VERSION : 0.1
   VAR_INPUT
      codeLib : "From Excel: Data";
   END_VAR
   VAR_IN_OUT
      savedWipStns : "Recipe: HMI Stations Saved Wips";
   END_VAR
   VAR_TEMP
      pStn : Int;
      pDestStn : Int;
      pWip : Int;
   END_VAR
BEGIN
   REGION "HMI STATIONS"
       FOR #pStn := 0 TO UDINT_TO_INT("Length"(#codeLib.hmiStns) - 1) DO
           #pDestStn := #codeLib.hmiStns[#pStn].pStn;
           IF #pDestStn = -1 THEN
               EXIT;
           END_IF;
           FOR #pWip := 0 TO "wipCount" DO
               #savedWipStns.stn[#pStn].wip[#pWip].pnCode :=
                   #codeLib.hmiStns[#pStn].wip[#pWip].pnCode;
           END_FOR;
       END_FOR;
   END_REGION
END_FUNCTION

FUNCTION "From Excel: PN Code to HMI Stations" : Void   // FC62, SCL
{ S7_Optimized_Access := 'TRUE' }
VERSION : 0.1
   VAR_INPUT
      xlCodeLib : "From Excel: Data";
   END_VAR
   VAR_IN_OUT
      stns : "Station: All Stations";
   END_VAR
   VAR_TEMP
      pSrc : Int;
      pDest : Int;
   END_VAR
BEGIN
   REGION "HMI STATIONS"
       FOR #pSrc := 0 TO UDINT_TO_INT("Length"(#xlCodeLib.hmiStns) - 1) DO
           #pDest := #xlCodeLib.hmiStns[#pSrc].pStn;
           IF #pDest = -1 THEN
               EXIT;
           END_IF;
           #stns.stn[#pDest].wipCmpts.pnCode := #xlCodeLib.hmiStns[#pSrc].wip[0].pnCode;
       END_FOR;
   END_REGION
END_FUNCTION

FUNCTION "From Excel: Wip Code to HMI Station Saved WIps" : Void   // FC63, SCL
{ S7_Optimized_Access := 'TRUE' }
VERSION : 0.1
   VAR_INPUT
      xlCodeLib : "From Excel: Data";
   END_VAR
   VAR_IN_OUT
      savedWipStns : "Recipe: HMI Stations Saved Wips";
   END_VAR
   VAR_TEMP
      pStn : Int;
      pDestStn : Int;
      pWip : Int;
   END_VAR
BEGIN
   REGION "HMI STATIONS"
       FOR #pStn := 0 TO UDINT_TO_INT("Length"(#xlCodeLib.hmiStns) - 1) DO
           FOR #pWip := 0 TO "wipCount" DO
               #savedWipStns.stn[#pStn].wip[#pWip].wip.code :=
                   #xlCodeLib.hmiStns[#pStn].wip[#pWip].wipCode;
           END_FOR;
       END_FOR;
   END_REGION
END_FUNCTION

// folder: Global/Physical

FUNCTION "Physical to Global" : Void   // FC1, LAD
{ S7_Optimized_Access := 'TRUE' }
VERSION : 0.1
   VAR_IN_OUT
      stations : "Station: All Stations";
   END_VAR
   VAR_TEMP
      i : Int;
      kp8In : DWord;
   END_VAR
BEGIN

REGION Network 1 (SCL): MAIN LOOP
   FOR #i := 0 TO "stnCount" DO

       CASE #i OF
           "VOLVO 16 01":
               #kp8In := "VOLVO 16 01 KP8 In";
           "VOLVO 16 02":
               #kp8In := "VOLVO 16 02 KP8 In";
           "VOLVO 16 03":
               #kp8In := "VOLVO 16 03 KP8 In";
           "VOLVO 16 04":
               #kp8In := "VOLVO 16 04 KP8 In";
           "VOLVO 16 05":
               #kp8In := "VOLVO 16 05 KP8 In";
           "VOLVO 16 06":
               #kp8In := "VOLVO 16 06 KP8 In";
           "VOLVO 16 07":
               #kp8In := "VOLVO 16 07 KP8 In";
           "VOLVO 16 08":
               #kp8In := "VOLVO 16 08 KP8 In";
           "VOLVO 16 09":
               #kp8In := "VOLVO 16 09 KP8 In";
           "VOLVO 16 10":
               #kp8In := "VOLVO 16 10 KP8 In";
           "VOLVO 16 11":
               #kp8In := "VOLVO 16 11 KP8 In";
           "CHM 01":
               #kp8In := "CHM 01 KP8 In";
           "CHM 02":
               #kp8In := "CHM 02 KP8 In";
           "CHM 03":
               #kp8In := "CHM 03 KP8 In";
           "CHM 04":
               #kp8In := "CHM 04 KP8 In";
           "CHM 05":
               #kp8In := "CHM 05 KP8 In";
           "CDO 01":
               #kp8In := "CDO 01 KP8 In";
           "CDO 02":
               #kp8In := "CDO 02 KP8 In";
           "CDO 03":
               #kp8In := "CDO 03 KP8 In";
           "BFL 01":
               #kp8In := "BFL 01 KP8 In";
           "BFL 02":
               #kp8In := "BFL 02 KP8 In";
           "BFL 03":
               #kp8In := "BFL 03 KP8 In";
           "LGS 01":
               #kp8In := "LGS 01 KP8 In";
           "LGS 02":
               #kp8In := "LGS 02 KP8 In";
           "LGS 03":
               #kp8In := "LGS 03 KP8 In";
           "CV 01":
               #kp8In := "CV 01 KP8 In";
           "CV 02":
               #kp8In := "CV 02 KP8 In";
           "CV 03":
               #kp8In := "CV 03 KP8 In";
           "CV 04":
               #kp8In := "CV 04 KP8 In";
           "PC 01":
               #kp8In := "PC 01 KP8 In"; 
           "PC 02":
               #kp8In := "PC 02 KP8 In";
       END_CASE;

       #stations.stn[#i].wipCmpts.ioData.kp8.input := #kp8In.%W1;

   END_FOR;
END_REGION
END_FUNCTION

FUNCTION "Global to Physical" : Void   // FC5, LAD
{ S7_Optimized_Access := 'TRUE' }
VERSION : 0.1
   VAR_IN_OUT
      stations : "Station: All Stations";
   END_VAR
   VAR_TEMP
      i : Int;
      j : Int;
      ET200SP : DWord;
      "KP8 In" : DWord;
      "KP8 Out" : DWord;
      Card : Int;
      stnCount : Int;
   END_VAR
BEGIN

REGION Network 1 (SCL): MAIN LOOP
   FOR #i := 0 TO "stnCount" DO

       #ET200SP := #stations.stn[#i].wipCmpts.ioData.stkLight;
       #"KP8 Out" := #stations.stn[#i].wipCmpts.ioData.kp8.tempOut;

       CASE #i OF
           "VOLVO 16 01":
               "VOLVO 16 01 IO" := #ET200SP;
               "VOLVO 16 01 KP8 Out" := #"KP8 Out";
           "VOLVO 16 02":
               "VOLVO 16 02 IO" := #ET200SP;
               "VOLVO 16 02 KP8 Out" := #"KP8 Out";
           "VOLVO 16 03":
               "VOLVO 16 03 IO" := #ET200SP;
               "VOLVO 16 03 KP8 Out" := #"KP8 Out";
           "VOLVO 16 04":
               "VOLVO 16 04 IO" := #ET200SP;
               "VOLVO 16 04 KP8 Out" := #"KP8 Out";
           "VOLVO 16 05":
               "VOLVO 16 05 IO" := #ET200SP;
               "VOLVO 16 05 KP8 Out" := #"KP8 Out";
           "VOLVO 16 06":
               "VOLVO 16 06 IO" := #ET200SP;
               "VOLVO 16 06 KP8 Out" := #"KP8 Out";
           "VOLVO 16 07":
               "VOLVO 16 07 IO" := #ET200SP;
               "VOLVO 16 07 KP8 Out" := #"KP8 Out";
           "VOLVO 16 08":
               "VOLVO 16 08 IO" := #ET200SP;
               "VOLVO 16 08 KP8 Out" := #"KP8 Out";
           "VOLVO 16 09":
               "VOLVO 16 09 IO" := #ET200SP;
               "VOLVO 16 09 KP8 Out" := #"KP8 Out";
           "VOLVO 16 10":
               "VOLVO 16 10 IO" := #ET200SP;
               "VOLVO 16 10 KP8 Out" := #"KP8 Out";
           "VOLVO 16 11":
               "VOLVO 16 11 IO" := #ET200SP;
               "VOLVO 16 11 KP8 Out" := #"KP8 Out";
           "CHM 01":
               "CHM 01 IO" := #ET200SP;
               "CHM 01 KP8 Out" := #"KP8 Out";
           "CHM 02":
               "CHM 02 IO" := #ET200SP;
               "CHM 02 KP8 Out" := #"KP8 Out";
           "CHM 03":
               "CHM 03 IO" := #ET200SP;
               "CHM 03 KP8 Out" := #"KP8 Out";
           "CHM 04":
               "CHM 04 IO" := #ET200SP;
               "CHM 04 KP8 Out" := #"KP8 Out";
           "CHM 05":
               "CHM 05 IO" := #ET200SP;
               "CHM 05 KP8 Out" := #"KP8 Out";
           "CDO 01":
               "CDO 01 IO" := #ET200SP;
               "CDO 01 KP8 Out" := #"KP8 Out";
           "CDO 02":
               "CDO 02 IO" := #ET200SP;
               "CDO 02 KP8 Out" := #"KP8 Out";
           "CDO 03":
               "CDO 03 IO" := #ET200SP;
               "CDO 03 KP8 Out" := #"KP8 Out";
           "BFL 01":
               "BFL 01 IO" := #ET200SP;
               "BFL 01 KP8 Out" := #"KP8 Out";
           "BFL 02":
               "BFL 02 IO" := #ET200SP;
               "BFL 02 KP8 Out" := #"KP8 Out";
           "BFL 03":
               "BFL 03 IO" := #ET200SP;
               "BFL 03 KP8 Out" := #"KP8 Out";
           "LGS 01":
               "LGS 01 IO" := #ET200SP;
               "LGS 01 KP8 Out" := #"KP8 Out";
           "LGS 02":
               "LGS 02 IO" := #ET200SP;
               "LGS 02 KP8 Out" := #"KP8 Out";
           "LGS 03":
               "LGS 03 IO" := #ET200SP;
               "LGS 03 KP8 Out" := #"KP8 Out";
           "CV 01":
               "CV 01 IO" := #ET200SP;
               "CV 01 KP8 Out" := #"KP8 Out";
           "CV 02":
               "CV 02 IO" := #ET200SP;
               "CV 02 KP8 Out" := #"KP8 Out";
           "CV 03":
               "CV 03 IO" := #ET200SP;
               "CV 03 KP8 Out" := #"KP8 Out";
           "CV 04":
               "CV 04 IO" := #ET200SP;
               "CV 04 KP8 Out" := #"KP8 Out";
           "PC 01":
               "PC 01 IO" := #ET200SP;
               "PC 01 KP8 Out" := #"KP8 Out";
           "PC 02":
               "PC 02 IO" := #ET200SP;
               "PC 02 KP8 Out" := #"KP8 Out";

       END_CASE;

   END_FOR;
END_REGION
END_FUNCTION

// folder: HMI: Warehouse/001 Part Call

FUNCTION_BLOCK "Part Call"   // FB16, SCL
{ S7_Optimized_Access := 'TRUE' }
VERSION : 0.1
   VAR_INPUT
      tblData : "Part Request Data";
      stns : "Station: All Stations";
      savedWips : "Recipe: HMI Stations Saved Wips";
      pnLib : "Recipe: PN Text Library";
   END_VAR
   VAR_IN_OUT
      tblHMI : "Part Call Screen";
      tableNav : "Nav Bar Data: PLC";
   END_VAR
   VAR RETAIN
      rowIndices : Array[0.."partReqTblHMIRowCnt"] of DInt;
   END_VAR
   VAR
      "inst Table Nav" : "Table Nav";
   END_VAR
   VAR_TEMP
      _tblHMI : "Part Call Screen";
      pRowHMI : DInt;
      pRowData : DInt;
   END_VAR
   // rowIndices[1] := 1;
   // rowIndices[2] := 2;
   // rowIndices[3] := 3;
   // rowIndices[4] := 4;
   // rowIndices[5] := 5;
   // rowIndices[6] := 6;
   // rowIndices[7] := 7;
   // rowIndices[8] := 8;
   // rowIndices[9] := 9;
   // rowIndices[10] := 10;
BEGIN
   REGION "TABLE NAVIGATION"
       #"inst Table Nav"(tblData := #tblData.row,
                         tblDisp := #tblHMI.row,
                         tableNav := #tableNav,
                         rowIndices := #rowIndices);
   END_REGION


   REGION "NAV BUTTON ANIMATIONS"
       "Part Call: Nav Animations"(#tableNav);
   END_REGION

   REGION "DOUBLE BUFFER IN"
       #_tblHMI := #tblHMI;
   END_REGION

   REGION "DRAW HMI TABLE"
       FOR #pRowHMI := 0 TO "partReqTblHMIRowCnt" DO

           REGION "ROW POINTER"
               #pRowData := #rowIndices[#pRowHMI];
           END_REGION

           REGION "DATA"
               "Part Call: Populate HMI Row"(address := #tblData.row[#pRowData],
                                             pnLib := #pnLib,
                                             stns := #stns,
                                             hmiRow := #_tblHMI.row[#pRowHMI]);
           END_REGION

           REGION "ANIMATIONS"
               "Part Call: Row Animations"(address := #tblData.row[#pRowData],
                                           stns := #stns,
                                           savedWips := #savedWips,
                                           rowHMI := #_tblHMI.row[#pRowHMI]);
           END_REGION

       END_FOR;
   END_REGION

   REGION "DOUBLE BUFFER OUT"
       #tblHMI := #_tblHMI;
   END_REGION
END_FUNCTION_BLOCK

FUNCTION "Part Call: Nav Animations" : Void   // FC18, SCL
{ S7_Optimized_Access := 'TRUE' }
VERSION : 0.1
   VAR_IN_OUT
      tableNav : "Nav Bar Data: PLC";
   END_VAR
   VAR_TEMP
      gray : USInt;
      green : USInt;
   END_VAR
BEGIN
   REGION "ANIMATE PART CALL NAV"

       REGION "COPY TO LOCAL"
           #gray := "BgGray";
           #green := "BgLGr";
       END_REGION

       REGION "TOP"
           #tableNav.top.animate := "Animate Bool"(colorTrue := #green,
                                                   colorFalse := #gray,
                                                   evalSignal := #tableNav.top.actuate);
       END_REGION

       REGION "PAGE UP"
           #tableNav.pageUp.animate := "Animate Bool"(colorTrue := #green,
                                                      colorFalse := #gray,
                                                      evalSignal := #tableNav.pageUp.actuate);
       END_REGION

       REGION "LINE UP"
           #tableNav.lineUp.animate := "Animate Bool"(colorTrue := #green,
                                                      colorFalse := #gray,
                                                      evalSignal := #tableNav.lineUp.actuate);
       END_REGION

       REGION "LINE DOWN"
           #tableNav.lineDown.animate := "Animate Bool"(colorTrue := #green,
                                                        colorFalse := #gray,
                                                        evalSignal := #tableNav.lineDown.actuate);
       END_REGION

       REGION "PAGE DOWN"
           #tableNav.pageDown.animate := "Animate Bool"(colorTrue := #green,
                                                        colorFalse := #gray,
                                                        evalSignal := #tableNav.pageDown.actuate);
       END_REGION

       REGION "BOTTOM"
           #tableNav.bottom.animate := "Animate Bool"(colorTrue := #green,
                                                      colorFalse := #gray,
                                                      evalSignal := #tableNav.bottom.actuate);
       END_REGION

   END_REGION
END_FUNCTION

FUNCTION "Part Call: Populate HMI Row" : Void   // FC19, SCL
{ S7_Optimized_Access := 'TRUE' }
VERSION : 0.1
   VAR_INPUT
      address : DInt;
      pnLib : "Recipe: PN Text Library";
      stns : "Station: All Stations";
   END_VAR
   VAR_IN_OUT
      hmiRow : "Table Row";
   END_VAR
   VAR_TEMP
      saveAct : Bool;
      pStn : DInt;
      pWip : DInt;
      pBtn : DInt;
      blankRow : "Table Row";
   END_VAR
BEGIN
   REGION "ROW HAS DATA"
       IF #address <> -1 THEN

           REGION "GET POINTERS"
               #pStn := "Address: Get Station"(#address);
               #pWip := "Address: Get Wip"(#address);
               #pBtn := "Address: Get Button"(#address);
           END_REGION

           REGION "NON WIP SPECIFIC"

           END_REGION

           REGION "GET DATA"
               #hmiRow.address := #address;
               #hmiRow.ordered := "Part Ordered"(#stns.stn[#pStn].wipCmpts.orderState[#pBtn]);
               #hmiRow.tfDropZone.value := "Strip Sign"(USINT_TO_WSTRING(#stns.stn[#pStn].id.dropZone));
               #hmiRow.tfLine.value := #stns.stn[#pStn].id.lineName;
               #hmiRow.tfPartNumber.value := "Get PN From Library"(pnLib := #pnLib, pnCode := #stns.stn[#pStn].wipCmpts.pnCode[#pBtn]);
               #hmiRow.tfTime.value := "Timer: Real to WString"(#stns.stn[#pStn].wipCmpts.timers.remaining[#pBtn]);
           END_REGION

       END_IF;
   END_REGION

   REGION "ROW HAS NO DATA"
       IF #address = -1 THEN
           #hmiRow := #blankRow;
       END_IF;
   END_REGION
END_FUNCTION

FUNCTION "Part Call: Row Animations" : Void   // FC20, SCL
{ S7_Optimized_Access := 'TRUE' }
VERSION : 0.1
   VAR_INPUT
      address : DInt;
      stns : "Station: All Stations";
      savedWips : "Recipe: HMI Stations Saved Wips";
   END_VAR
   VAR_IN_OUT
      rowHMI : "Table Row";
   END_VAR
   VAR_TEMP
      cBackground : USInt;
      cForeground : USInt;
      state : Int;
   END_VAR
BEGIN
   REGION "ROW HAS DATA"
       IF #address >= 0 THEN

           REGION "GET STATE"
               #state := "Part Call: Get State"(address := #address,
                                                stns := #stns,
                                                savedWips := #savedWips);
           END_REGION

           REGION "GET COLOR"
               "Part Call: State to Color"(state := #state,
                                           background => #cBackground,
                                           foreground => #cForeground);
           END_REGION

       END_IF;
   END_REGION

   REGION "ROW HAS NO DATA"
       IF #address <= -1 THEN
           #cForeground := "invisible";
           #cBackground := "invisible";
       END_IF;
   END_REGION


   REGION "DRAW TO HMI"
       "Part Call: Color Row"(cBackground := #cBackground,
                              cForeground := #cForeground,
                              singleLinePN := TRUE,
                              rowHMI := #rowHMI);
   END_REGION
END_FUNCTION

FUNCTION "Part Call: State to Color" : Void   // FC22, SCL
{ S7_Optimized_Access := 'TRUE' }
VERSION : 0.1
   VAR_INPUT
      state : Int;
   END_VAR
   VAR_OUTPUT
      background : USInt;
      foreground : USInt;
   END_VAR
   VAR_TEMP
      bg : USInt;
      cBlue : USInt;
      cGrayLight : USInt;
      cGrayDark : USInt;
      cGreen : USInt;
      cInvisible : USInt;
      cRedSolid : USInt;
      cRedFlash : USInt;
      cWhite : USInt;
      fg : USInt;
   END_VAR
BEGIN
   #cBlue := "BgLBl";
   #cGreen := "BgLGr";
   #cInvisible := "invisible";
   #cRedSolid := "BgLRd";
   #cRedFlash := "FlLRd";
   #cGrayLight := "BgGray";
   #cGrayDark := "disabled";
   #cWhite := "BgWh";

   CASE #state OF
       0, "idle":
           #bg := #cInvisible;
           #fg := #cInvisible;
       "requested", "acknowledged":
           #bg := #cGrayDark;
           #fg := #cGrayLight;
       "requestedCrit", "orderedCrit", "acknowledgedCrit":
           #bg := #cGrayDark;
           #fg := #cRedSolid;
       "requestedExp", "orderedExp", "acknowledgedExp":
           #bg := #cGrayDark;
           #fg := #cRedFlash;
       "ordered":
           #bg := #cGrayDark;
           #fg := #cBlue;
   END_CASE;

   #foreground := #fg;
   #background := #bg;
END_FUNCTION

FUNCTION "Part Call: Color Row" : Void   // FC31, SCL
{ S7_Optimized_Access := 'TRUE' }
VERSION : 0.1
   VAR_INPUT
      cBackground : USInt;
      cForeground : USInt;
      singleLinePN : Bool;
   END_VAR
   VAR_IN_OUT
      rowHMI : "Table Row";
   END_VAR
   VAR_TEMP
      row : "Table Row";
   END_VAR
BEGIN
   REGION "DOUBLE BUFFER IN"
       #row := #rowHMI;
   END_REGION

   REGION "INDEPENDANT ROWS"
       #row.pbSelection.animate := #cForeground;
       #row.rtBackground.animate := #cBackground;
       #row.tfDropZone.animate := #cForeground;
       #row.tfLine.animate := #cForeground;
       #row.tfTime.animate := #cForeground;
   END_REGION


   REGION "DEPENDANT ROWS"

       REGION "SINGLE LINE PART NUMBER"
           IF #singleLinePN THEN
               #row.tfPartNumber.animateDL := "invisible";
               #row.tfPartNumber.animateSL := #cForeground;
           END_IF;
       END_REGION

       REGION "DOUBLE LINE PN"
           IF NOT #singleLinePN THEN
               #row.tfPartNumber.animateDL := #cForeground;
               #row.tfPartNumber.animateSL := "invisible";
           END_IF;
       END_REGION

   END_REGION

   REGION "DOUBLE BUFFER OUT"
       #rowHMI := #row;
   END_REGION
END_FUNCTION

FUNCTION "Address in Loaded Wip" : Bool   // FC43, SCL
{ S7_Optimized_Access := 'TRUE' }
VERSION : 0.1
   VAR_INPUT
      pWip : DInt;
      stn : "Station: Single Station";
   END_VAR
   VAR_TEMP
      ret : Bool;
   END_VAR
BEGIN
   IF #pWip = #stn.wipData.index THEN
       #ret := TRUE;
   END_IF;
   #"Address in Loaded Wip" := #ret;
END_FUNCTION

FUNCTION "Part Call: Get State" : Int   // FC57, SCL
{ S7_Optimized_Access := 'TRUE' }
VERSION : 0.1
   VAR_INPUT
      address : DInt;
      stns : "Station: All Stations";
      savedWips : "Recipe: HMI Stations Saved Wips";
   END_VAR
   VAR_TEMP
      addressInWip : Bool;
      pBtn : DInt;
      pStn : DInt;
      pWip : DInt;
      ret : Int;
   END_VAR
BEGIN
   REGION "DECOMPOSE ADDRESS"
       #pBtn := "Address: Get Button"(#address);
       #pStn := "Address: Get Station"(#address);
       #pWip := "Address: Get Wip"(#address);
   END_REGION

   REGION "CHECK ADDRESS AGAINST STATION'S CURRENT WIP"
       #addressInWip := "Address in Loaded Wip"(pWip := #pWip,
                                                stn := #stns.stn[#pStn]);
   END_REGION

   REGION "ADDRESS IN WIP"
       IF #addressInWip THEN
           #ret := #stns.stn[#pStn].wipCmpts.orderState[#pBtn];
       END_IF;
   END_REGION

   REGION "ADDRESS NOT IN WIP"
       IF NOT #addressInWip THEN
           #ret := #savedWips.stn[#pStn].wip[#pWip].orderState[#pBtn];
       END_IF;
   END_REGION

   REGION "RETURN"
       #"Part Call: Get State" := #ret;
   END_REGION
END_FUNCTION

// folder: HMI: Warehouse/002 Settings

FUNCTION_BLOCK "Settings Screen"   // FB19, SCL
{ S7_Optimized_Access := 'TRUE' }
VERSION : 0.1
   VAR_INPUT
      selected_stations : "Selected Stations";
      selected_buttons : "Selected Buttons";
      selected_wips : "Selected Wips";
      stations : "Station: All Stations";
   END_VAR
   VAR_IN_OUT
      settings : "Settings";
   END_VAR
   VAR
      "Table Nav_Instance" : "Table Nav";
   END_VAR
BEGIN
   REGION "ANIMATION"
       "Settings Screen: Animations"(selected_stations := #selected_stations,
                                     selected_buttons := #selected_buttons,
                                     selected_wips := #selected_wips,
                                     stations := #stations,
                                     screen := #settings);
   END_REGION
END_FUNCTION_BLOCK

FUNCTION "Settings Screen: Animations: Select Stations Button" : Void   // FC92, SCL
{ S7_Optimized_Access := 'TRUE' }
VERSION : 0.1
   VAR_IN_OUT
      interface : "PB Data";
   END_VAR
   VAR_TEMP
      t_interface : "PB Data";
   END_VAR
BEGIN
   REGION "COPY TO LOCAL"
       #t_interface := #interface;
   END_REGION


   REGION "ANIMATE"
       #t_interface.animate := "Animate Bool"(colorTrue := "BgLGr",
                                              colorFalse := "BgGray",
                                              evalSignal := #t_interface.actuate);
       #t_interface.enable := TRUE;
       #t_interface.visible := TRUE;
   END_REGION


   REGION "DRAW"
       #interface := #t_interface;
   END_REGION
END_FUNCTION

FUNCTION "Settings Screen: Animations: Select WIP Button" : Void   // FC93, SCL
{ S7_Optimized_Access := 'TRUE' }
VERSION : 0.1
   VAR_INPUT
      selected_stations : "Selected Stations";
      stations : "Station: All Stations";
   END_VAR
   VAR_IN_OUT
      select_wip : "PB Data";
   END_VAR
   VAR_TEMP
      index_of_first_selected_station : Int;
      is_hmi_station : Bool;
      first_selected_station : "Station: Single Station";
      t_select_wip : "PB Data";
   END_VAR
BEGIN
   REGION "COPY TO LOCAL"
       #t_select_wip := #select_wip;
   END_REGION

   REGION "ARE SELECTED STATIONS HMI STATIONS?"
       #index_of_first_selected_station := "Get First Selected Station"(#selected_stations.stns);
       #first_selected_station := #stations.stn[#index_of_first_selected_station];
       #is_hmi_station := "Is HMI Station"(#first_selected_station);
   END_REGION

   REGION "HMI STATIONS"
       IF #is_hmi_station THEN
           #t_select_wip.animate := "Animate Bool"(colorTrue := "BgLGr",
                                                   colorFalse := "BgGray",
                                                   evalSignal := #t_select_wip.actuate);
           #t_select_wip.enable := TRUE;
           #t_select_wip.visible := TRUE;
       END_IF;
   END_REGION

   REGION "NON-HMI STATIONS"
       IF NOT #is_hmi_station THEN
           #t_select_wip.enable := FALSE;
           #t_select_wip.visible := FALSE;
       END_IF;
   END_REGION

   REGION "DRAW" 
       #select_wip := #t_select_wip;
   END_REGION
END_FUNCTION

FUNCTION "Settings Screen: Animations: Select Buttons Button" : Void   // FC94, SCL
{ S7_Optimized_Access := 'TRUE' }
VERSION : 0.1
   VAR_IN_OUT
      selectButton : "PB Data";
   END_VAR
   VAR_TEMP
      ret : "PB Data";
   END_VAR
BEGIN
   REGION "BUTTON ON"
       IF #selectButton.actuate THEN
           #ret.animate := "FgLGr";
       END_IF;
   END_REGION


   REGION "BUTTON OFF"
       IF NOT #selectButton.actuate THEN
           #ret.animate := "FgGray";
       END_IF;
   END_REGION


   REGION "DOUBLE BUFFER"
       #selectButton := #ret;
   END_REGION ;
END_FUNCTION

FUNCTION "Settings Screen: Animations" : Void   // FC123, SCL
{ S7_Optimized_Access := 'TRUE' }
VERSION : 0.1
   VAR_INPUT
      selected_stations : "Selected Stations";
      selected_buttons : "Selected Buttons";
      selected_wips : "Selected Wips";
      stations : "Station: All Stations";
   END_VAR
   VAR_IN_OUT
      screen : "Settings";
   END_VAR
   VAR_TEMP
      t_screen : "Settings";
   END_VAR
BEGIN
   REGION "COPY TO LOCAL"
       #t_screen := #screen;
   END_REGION


   REGION "SELECT STATION BUTTON ANIMATION"
       "Settings Screen: Animations: Select Stations Button"(#t_screen.selectStation);
   END_REGION


   REGION "SELECT BUTTONS BUTTON ANIMATION"    
   END_REGION


   REGION "SELECT WIP BUTTON ANIMATION"
       "Settings Screen: Animations: Select WIP Button"(selected_stations := #selected_stations,
                                                        stations := #stations,
                                                        select_wip := #t_screen.selectWip);
   END_REGION

   REGION "ASSIGN BUTTON ANIMATION"
       "Settings Screen: Animations: Assign Button"(selected_stations := #selected_stations,
                                                    selected_buttons := #selected_buttons,
                                                    selected_wips := #selected_wips,
                                                    stations := #stations,
                                                    interface := #t_screen.assign);
   END_REGION


   REGION "DRAW"
       #screen := #t_screen;
   END_REGION
END_FUNCTION

FUNCTION "Settings Screen: Animations: Assign Button" : Void   // FC124, SCL
{ S7_Optimized_Access := 'TRUE' }
VERSION : 0.1
   VAR_INPUT
      selected_stations : "Selected Stations";
      selected_buttons : "Selected Buttons";
      selected_wips : "Selected Wips";
      stations : "Station: All Stations";
   END_VAR
   VAR_IN_OUT
      interface : "PB Data";
   END_VAR
   VAR_TEMP
      enable : Bool;
      is_hmi_station : Bool;
      selected_stations_count : Int;
      selected_buttons_count : Int;
      selected_wips_count : Int;
      t_interface : "PB Data";
      visible : Bool;
   END_VAR
BEGIN
   REGION "COPY TO LOCAL"
       #t_interface := #interface;
   END_REGION


   REGION "GET COUNTS"
       #selected_stations_count := "Count Selected Stations"(#selected_stations.stns);
       #selected_buttons_count := "Count Selected Buttons"(#selected_buttons.btns);
       #selected_wips_count := "Count Selected WIPs"(#selected_wips.wips);
   END_REGION


   REGION "STATIONS ARE HMI STATIONS"
       #is_hmi_station := "Is HMI Station"(#stations.stn["Get First Selected Station"(#selected_stations.stns)]);
   END_REGION


   REGION "ENABLE AND MAKE VISIBLE"
       IF (#selected_buttons_count > 0) AND
           (#selected_stations_count > 0) AND
           ((#is_hmi_station AND #selected_wips_count > 0) OR NOT #is_hmi_station) THEN
               #enable := TRUE;
               #visible := TRUE;
       END_IF;
   END_REGION


   REGION "ANIMATION"
       IF #enable AND #visible THEN
           #t_interface.animate := "Animate Bool"(colorTrue := "BgLGr",
                                                  colorFalse := "BgGray",
                                                  evalSignal := #t_interface.actuate);
       END_IF;
   END_REGION


   REGION "ENABLE"
       #t_interface.enable := #enable;
   END_REGION


   REGION "VISIBLE"
       #t_interface.visible := #visible;
   END_REGION


   REGION "DRAW" 
       #interface := #t_interface;
   END_REGION
END_FUNCTION

// folder: HMI: Warehouse/Pop Ups/Pop Up Utilities

FUNCTION "Pop Up: Map Select Button Actuations" : Void   // FC117, SCL
{ S7_Optimized_Access := 'TRUE' }
VERSION : 0.1
   VAR_INPUT
      screen_elements : Variant;
   END_VAR
   VAR_IN_OUT
      actuations_as_ints : Variant;
   END_VAR
   VAR_TEMP
      i : Int;
      len_udint : UDInt;
      len_int : Int;
      ret : Array[0..#u_bound] of Int;
      status : Int;
      t_select_btns : Array[0..#u_bound] of "PB Data";
   END_VAR
   VAR CONSTANT
      u_bound : Int := 99;
   END_VAR
BEGIN
   #len_udint := CountOfElements(#screen_elements);
   #len_int := UDINT_TO_INT(#len_udint) - 1;
   #status := MOVE_BLK_VARIANT(SRC := #screen_elements,
                               COUNT := #len_udint,
                               SRC_INDEX := 0,
                               DEST_INDEX := 0,
                               DEST => #t_select_btns);
   FOR #i := 0 TO #len_int DO
       IF #t_select_btns[#i].actuate THEN
           #ret[#i] := 1;
       END_IF;
   END_FOR;
   #status := MOVE_BLK_VARIANT(SRC := #ret,
                               COUNT := #len_udint,
                               SRC_INDEX := 0,
                               DEST_INDEX := 0,
                               DEST => #actuations_as_ints);
END_FUNCTION

// folder: HMI: Warehouse/Pop Ups/Select Buttons

FUNCTION_BLOCK "Pop Up: Select Buttons"   // FB25, SCL
{ S7_Optimized_Access := 'TRUE' }
VERSION : 0.1
   VAR_IN_OUT
      interface : "Select Button";
      selected_buttons : "Selected Buttons";
   END_VAR
   VAR
      "inst Pop Up: Select Buttons: Select Buttons" : "Pop Up: Select Buttons: Select Buttons";
   END_VAR
BEGIN
   REGION "ANIMATION"
       "Pop Up: Select Buttons: Animations"(interface := #interface,
                                            selected := #selected_buttons);
   END_REGION


   REGION "PERFORM BUTTON SELECTION"
       #"inst Pop Up: Select Buttons: Select Buttons"(interface := #interface,
                                                      selected_buttons := #selected_buttons);
   END_REGION
END_FUNCTION_BLOCK

FUNCTION_BLOCK "Pop Up: Select Buttons: Select Buttons"   // FB27, SCL
{ S7_Optimized_Access := 'TRUE' }
VERSION : 0.1
   VAR_IN_OUT
      interface : "Select Button";
      selected_buttons : "Selected Buttons";
   END_VAR
   VAR
      "inst Pulses: Button Collection" : "Pulses: Button Collection";
   END_VAR
   VAR_TEMP
      actuation_pulses : Array[0.."btnCount"] of Bool;
      actuations_as_ints : Array[0.."btnCount"] of Int;
      i : Int;
      pulses_as_ints : Array[0.."btnCount"] of Int;
   END_VAR
BEGIN
   "Pop Up: Map Select Button Actuations"(screen_elements := #interface.buttons,
                                          actuations_as_ints := #actuations_as_ints);
   #"inst Pulses: Button Collection"(btns := #actuations_as_ints,
                                     pulses := #pulses_as_ints);
   "Pop Up: Select Buttons: Pulse Ints to Bools"(pulses_as_ints := #pulses_as_ints,
                                                 pulses_as_bools => #actuation_pulses);
   FOR #i := 0 TO "btnCount" DO
       "Toggle"(pulse := #actuation_pulses[#i],
                state := #selected_buttons.btns[#i]);
   END_FOR;
END_FUNCTION_BLOCK

FUNCTION "Pop Up: Select Buttons: Animations" : Void   // FC116, SCL
{ S7_Optimized_Access := 'TRUE' }
VERSION : 0.1
   VAR_IN_OUT
      interface : "Select Button";
      selected : "Selected Buttons";
   END_VAR
   VAR_TEMP
      i : Int;
      selected_stations_count : Int;
      t_interface : "Select Button";
   END_VAR
BEGIN
   REGION "COPY TO LOCAL"
       #t_interface := #interface;
   END_REGION

   REGION "CLOSE POPUP BUTTON"
       #t_interface.close_screen.animate := "Animate Bool"(colorTrue := "BgLGr",
                                                           colorFalse := "BgLRd",
                                                           evalSignal := #interface.close_screen.actuate);
   END_REGION


   REGION "BUTTON SELECTION BUTTONS"
       FOR #i := 0 TO "btnCount" DO
           #t_interface.buttons[#i].animate := "Animate Bool"(colorTrue := "BgLGr",
                                                              colorFalse := "BgGray",
                                                              evalSignal := #interface.buttons[#i].actuate);
           #t_interface.buttons[#i].enable := TRUE;
           #t_interface.buttons[#i].visible := TRUE;
           IF #selected.btns[#i] THEN
               #t_interface.buttons[#i].animate := "BgLBl";
           END_IF;
       END_FOR;
   END_REGION


   REGION "DRAW"
       #interface := #t_interface;
   END_REGION
END_FUNCTION

FUNCTION "Pop Up: Select Buttons: Pulse Ints to Bools" : Void   // FC118, SCL
{ S7_Optimized_Access := 'TRUE' }
VERSION : 0.1
   VAR_INPUT
      pulses_as_ints : Array[0.."btnCount"] of Int;
   END_VAR
   VAR_OUTPUT
      pulses_as_bools : Array[0.."btnCount"] of Bool;
   END_VAR
   VAR_TEMP
      i : Int;
      ret : Array[0.."btnCount"] of Bool;
   END_VAR
BEGIN
   REGION "MAP TO BOOLS"
       FOR #i := 0 TO "btnCount" DO
           #ret[#i] := #pulses_as_ints[#i].%X0;
       END_FOR;
   END_REGION

   REGION "RETURN"
       #pulses_as_bools := #ret;
   END_REGION
END_FUNCTION

// folder: HMI: Warehouse/Pop Ups/Select Station

FUNCTION_BLOCK "Pop Up: Select Stations"   // FB21, SCL
{ S7_Optimized_Access := 'TRUE' }
VERSION : 0.1
   VAR_IN_OUT
      all_stations : "Station: All Stations";
      interface : "Select Station";
      meta_data : "Setting Meta Data";
   END_VAR
   VAR
      "inst Patch for Table Nav in Select Station Popup" : "Patch for Table Nav in Select Station Popup";
      "inst Select Station Button Pulses" : "Pulses: Button Collection";
      "inst Selection Change" : "Pop Up: Select Stations: Selection Change";
      "inst Table Nav" : "Table Nav";
      selectable_stn_cnt : Int;
      vis_stns_as_dint : Array[0.."slct_stn_btn_count"] of DInt;
      visable_stns : Array[0.."slct_stn_btn_count"] of Int;
   END_VAR
   VAR_TEMP
      blank_station : "Station: Single Station";
      i : Int;
      nav_pulses : Int;
      p_stn : DInt;
      pulses_as_int : Array[0.."slct_stn_btn_count"] of Int;
      selectable_stns_as_dint : Array[0.."stnCount"] of DInt;
      selected_stn_cnt : Int;
      actuation_pulses : Array[0.."slct_stn_btn_count"] of Bool;
      actuations_as_ints : Array[0.."slct_stn_btn_count"] of Int;
      t_selection_change : "Station Selection Change";
   END_VAR
   // visable_stns[0] := 0;
   // visable_stns[1] := 1;
   // visable_stns[2] := 2;
   // visable_stns[3] := 3;
   // visable_stns[4] := 4;
   // visable_stns[5] := 5;
   // visable_stns[6] := 6;
   // visable_stns[7] := 7;
   // visable_stns[8] := 8;
   // visable_stns[9] := 9;
   // visable_stns[10] := 10;
   // visable_stns[11] := 11;
BEGIN
   REGION "ANIMATIONS"
       "Pop Up: Select Stations: Animations"(all_stations := #all_stations,
                                             selectable_stn_cnt := #selectable_stn_cnt,
                                             selected_stns := #meta_data.selected_stns,
                                             visable_stns := #visable_stns,
                                             interface := #interface);
   END_REGION


   REGION "CLEAR SELECTION CHANGE"
       #meta_data.selection_change := #t_selection_change;
   END_REGION


   REGION "SELECT STATION BUTTON PULSES"
       "Pop Up: Map Select Button Actuations"(screen_elements := #interface.stn_select_btns,
                                              actuations_as_ints := #actuations_as_ints);
       #"inst Select Station Button Pulses"(btns := #actuations_as_ints,
                                            pulses := #pulses_as_int);
       "Pop Up: Select Stations: Pulse Ints to Bools"(pulses_as_ints := #pulses_as_int,
                                                      pulses_as_bools => #actuation_pulses);
   END_REGION


   REGION "PERFORM STATION SELECTION"
       FOR #i := 0 TO "slct_stn_btn_count" DO
           IF #visable_stns[#i] <> -1 THEN
               "Toggle"(pulse := #actuation_pulses[#i],
                        state := #meta_data.selected_stns.stns[#visable_stns[#i]]);
           END_IF;
       END_FOR;
   END_REGION


   REGION "SCAN FOR CHANGE TO STATION SELECTION"
       #"inst Selection Change"(selected_stns := #meta_data.#selected_stns,
                                station_change => #meta_data.selection_change);
   END_REGION


   REGION "BUILD SELECTABLE STATION LIST"
       IF #meta_data.selection_change.selection_change OR "FirstScan" THEN
           "Build Selectable Station List"(selected_stns := #meta_data.selected_stns,
                                           selection_change := #meta_data.selection_change,
                                           stns := #all_stations,
                                           selectable_stns := #meta_data.selectable_stns.stns,
                                           visible_stations := #visable_stns,
                                           selectable_stn_cnt := #selectable_stn_cnt);
       END_IF;
   END_REGION


   REGION "TABLE NAV"

       // when there are more selectable stations than buttons
       IF #selectable_stn_cnt > "slct_stn_btn_count" THEN
           #"inst Table Nav"(first_null_index := #selectable_stn_cnt,
                             tblData := #selectable_stns_as_dint,
                             tblDisp := #vis_stns_as_dint,
                             tableNav := #interface.nav_Bar_PLC,
                             rowIndices := #vis_stns_as_dint);
           // patch for table nav to work with selectable stations
           #"inst Patch for Table Nav in Select Station Popup"(nav_bar := #interface.nav_Bar_PLC,
                                                               selectable_staions := #meta_data.selectable_stns.stns,
                                                               selection_change := #meta_data.selection_change.selection_change,
                                                               vis_stns_as_dint := #vis_stns_as_dint,
                                                               visable_stns := #visable_stns);
       END_IF;

       // when there are fewer selectable stations than buttons
       IF #selectable_stn_cnt < "slct_stn_btn_count" THEN
           IF #meta_data.selection_change.rising THEN
               "Fill Int Array"(int_in := -1,
                                array_out => #visable_stns);
               FOR #i := 0 TO #selectable_stn_cnt - 1 DO
                   #visable_stns[#i] := #meta_data.selectable_stns.stns[#i];
               END_FOR;
           END_IF;
       END_IF;


   END_REGION
END_FUNCTION_BLOCK

FUNCTION_BLOCK "Pop Up: Select Stations: Selection Change"   // FB23, SCL
{ S7_Optimized_Access := 'TRUE' }
VERSION : 0.1
   VAR_INPUT
      selected_stns : "Selected Stations";
   END_VAR
   VAR_OUTPUT
      station_change : "Station Selection Change";
   END_VAR
   VAR
      old : Struct
         selected_stns : "Selected Stations";
      END_STRUCT;
   END_VAR
   VAR_TEMP
      i : Int;
      ret : "Station Selection Change";
   END_VAR
BEGIN
   REGION "SCAN FOR CHANGE"
       FOR #i := 0 TO "stnCount" DO
           IF #selected_stns.stns[#i] <> #old.selected_stns.stns[#i] THEN
               #ret.selection_change := TRUE;
               #ret.station_index := #i;
               IF #selected_stns.stns[#i] AND NOT #old.selected_stns.stns[#i] THEN
                   #ret.rising := TRUE;
                   #ret.falling := FALSE;
               END_IF;
               IF NOT #selected_stns.stns[#i] AND #old.selected_stns.stns[#i] THEN
                   #ret.rising := FALSE;
                   #ret.falling := TRUE;
               END_IF;
               EXIT;
           END_IF;
       END_FOR;
   END_REGION


   REGION "SAVE TO OLD"
       #old.selected_stns := #selected_stns;
   END_REGION


   REGION "RETURN"
       #station_change.falling := #ret.falling;
       #station_change.rising := #ret.rising;
       #station_change.selection_change := #ret.selection_change;
       #station_change.station_index := #ret.station_index;
   END_REGION
END_FUNCTION_BLOCK

FUNCTION_BLOCK "Patch for Table Nav in Select Station Popup"   // FB24, SCL
{ S7_Optimized_Access := 'TRUE' }
VERSION : 0.1
   VAR_INPUT
      nav_bar : "Nav Bar Data: PLC";
      selectable_staions : Array[0.."stnCount"] of Int;
      selection_change : Bool;
   END_VAR
   VAR_IN_OUT
      vis_stns_as_dint : Array[0.."slct_stn_btn_count"] of DInt;
      visable_stns : Array[0.."slct_stn_btn_count"] of Int;
   END_VAR
   VAR
      old_nav : "Nav Bar Data: PLC";
   END_VAR
   VAR_TEMP
      i : Int;
      itrnl_visible_stns : Array[0.."slct_stn_btn_count"] of Int;
      nav_pulse : Bool;
      p_stn : DInt;
   END_VAR
BEGIN
   REGION "PULSE FROM ANY NAV BUTTON"
       IF NOT #old_nav.top.actuate AND #nav_bar.top.actuate THEN
           #nav_pulse := TRUE;
       END_IF;
       IF NOT #old_nav.pageUp.actuate AND #nav_bar.pageUp.actuate THEN
           #nav_pulse := TRUE;
       END_IF;
       IF NOT #old_nav.lineUp.actuate AND #nav_bar.lineUp.actuate THEN
           #nav_pulse := TRUE;
       END_IF;
       IF NOT #old_nav.lineDown.actuate AND #nav_bar.lineDown.actuate THEN
           #nav_pulse := TRUE;
       END_IF;
       IF NOT #old_nav.pageDown.actuate AND #nav_bar.pageDown.actuate THEN
           #nav_pulse := TRUE;
       END_IF;
       IF NOT #old_nav.bottom.actuate AND #nav_bar.bottom.actuate THEN
           #nav_pulse := TRUE;
       END_IF;
   END_REGION


   REGION "REMAP VISIBLE STATIONS BASED ON SELECTABLE STATIONS"
       IF #nav_pulse OR #selection_change THEN
           FOR #i := 0 TO "slct_stn_btn_count" DO
               #visable_stns[#i] := DINT_TO_INT(#vis_stns_as_dint[#i]);
               #itrnl_visible_stns[#i] := #selectable_staions[#visable_stns[#i]];
               #vis_stns_as_dint[#i] := INT_TO_DINT(#visable_stns[#i]);
           END_FOR;
           #visable_stns := #itrnl_visible_stns;
       END_IF;
   END_REGION


   REGION "SAVE FOR CHANGE DETECTION"
       #old_nav := #nav_bar;
   END_REGION
END_FUNCTION_BLOCK

FUNCTION "Select Station Button Activation" : Bool   // FC95, SCL
{ S7_Optimized_Access := 'TRUE' }
VERSION : 0.1
   VAR_INPUT
      btn_index : Int;
      selectable_stn_cnt : Int;
   END_VAR
   VAR_TEMP
      ret : Bool;
   END_VAR
BEGIN
   REGION "TURN ON A NUMBER OF BUTTONS EQUAL TO THE NUMBER OF STATIONS"
       IF #btn_index < #selectable_stn_cnt THEN
           #ret := TRUE;
       END_IF;
       IF #btn_index >= #selectable_stn_cnt THEN
           #ret := FALSE;
       END_IF;
   END_REGION

   REGION "RETURN"
       #"Select Station Button Activation" := #ret;
   END_REGION
END_FUNCTION

FUNCTION "Select Station Nav Bar Button Animation" : Void   // FC97, SCL
{ S7_Optimized_Access := 'TRUE' }
VERSION : 0.1
   VAR_INPUT
      selectable_stations : Int;
      visible_rows : Int;
   END_VAR
   VAR_IN_OUT
      button : "PB Data";
   END_VAR
   VAR_TEMP
      ret : "PB Data";
   END_VAR
BEGIN
   REGION "SHOW NAV BAR"
       IF #selectable_stations > #visible_rows THEN

           REGION "GET CURRENT STATE FOR PRESS"
               #ret := #button;
           END_REGION

           REGION "ANIMATION"
               #ret.animate := "Animate Bool"(colorTrue := "BgLGr",
                                              colorFalse := "BgGray",
                                              evalSignal := #button.actuate);
           END_REGION

           REGION "ENABLE"
               #ret.enable := TRUE;
           END_REGION

           REGION "LIST SELECT"
               #ret.listSelect := 0;
           END_REGION

           REGION "VISIBLE"
               #ret.visible := TRUE;
           END_REGION

       END_IF;
   END_REGION


   REGION "HIDE NAV BAR"
       IF #selectable_stations <= #visible_rows THEN

           REGION "DIABLE"
               #ret.enable := FALSE;
           END_REGION

           REGION "INVISIBLE"
               #ret.visible := FALSE;
           END_REGION

       END_IF;
   END_REGION


   REGION "RETURN"
       #button := #ret;
   END_REGION
END_FUNCTION

FUNCTION "Populate Station Name" : WString   // FC100, SCL
{ S7_Optimized_Access := 'TRUE' }
VERSION : 0.1
   VAR_INPUT
      lines : Int;
      stn : "Station: Single Station";
   END_VAR
   VAR_TEMP
      ret : WString;
      dz : WString;
   END_VAR
   VAR CONSTANT
      line_feed : WString := WSTRING#'$L';
   END_VAR
BEGIN
   REGION "FORMAT STRING"
       #dz := "Strip Sign"(USINT_TO_WSTRING(#stn.id.dropZone));
       #dz := "Add Leading"("Leading Character" := wchar#'0',
                            "Desired Length" := 2,
                            "String" := #dz);
   END_REGION

   REGION "ONE LINE"
       IF #lines = 1 THEN
           #ret := CONCAT_WSTRING(IN1 := #stn.id.lineName,
                                  IN2 := #dz);
       END_IF;
   END_REGION


   REGION "MORE THAN ONE LINE"
       IF #lines > 1 THEN
           #ret := CONCAT_WSTRING(IN1 := #stn.id.lineName,
                                  IN2 := #line_feed,
                                  IN3 := #dz);
       END_IF;
   END_REGION


   REGION "INVALID ENTRY"
       IF #lines < 1 THEN
           #ret := WString#'invalid line count';
       END_IF;
   END_REGION


   #"Populate Station Name" := #ret;
END_FUNCTION

FUNCTION "Pop Up: Select Stations: Map Select Button Acutations" : Void   // FC101, SCL
{ S7_Optimized_Access := 'TRUE' }
VERSION : 0.1
   VAR_INPUT
      select_btns : Array[0.."slct_stn_btn_count"] of "PB Data";
   END_VAR
   VAR_OUTPUT
      btn_actuations : Array[0.."slct_stn_btn_count"] of Int;
   END_VAR
   VAR_TEMP
      i : Int;
      ret : Array[0.."slct_stn_btn_count"] of Int;
   END_VAR
BEGIN
   REGION "MAP ACTUATIONS"
       FOR #i := 0 TO "slct_stn_btn_count" DO
           IF #select_btns[#i].actuate THEN
               #ret[#i] := 1;
           END_IF;
       END_FOR;
   END_REGION


   REGION "RETURN"
       #btn_actuations := #ret;
   END_REGION
END_FUNCTION

FUNCTION "Pop Up: Select Stations: Pulse Ints to Bools" : Void   // FC102, SCL
{ S7_Optimized_Access := 'TRUE' }
VERSION : 0.1
   VAR_INPUT
      pulses_as_ints : Array[0.."slct_stn_btn_count"] of Int;
   END_VAR
   VAR_OUTPUT
      pulses_as_bools : Array[0.."slct_stn_btn_count"] of Bool;
   END_VAR
   VAR_TEMP
      i : Int;
      ret : Array[0.."slct_stn_btn_count"] of Bool;
   END_VAR
BEGIN
   REGION "MAP TO BOOLS"
       FOR #i := 0 TO "slct_stn_btn_count" DO
           #ret[#i] := #pulses_as_ints[#i].%X0;
       END_FOR;
   END_REGION

   REGION "RETURN"
       #pulses_as_bools := #ret;
   END_REGION
END_FUNCTION

FUNCTION "Build Selectable Station List" : Void   // FC104, SCL
{ S7_Optimized_Access := 'TRUE' }
VERSION : 0.1
   VAR_INPUT
      selected_stns : "Selected Stations";
      selection_change : "Station Selection Change";
      stns : "Station: All Stations";
   END_VAR
   VAR_IN_OUT
      selectable_stns : Array[0.."stnCount"] of Int;
      visible_stations : Array[0.."slct_stn_btn_count"] of Int;
      selectable_stn_cnt : Int;
   END_VAR
   VAR_TEMP
      blank_stn : "Station: Single Station";
      eval_station_is_hmi : Bool;
      i : Int;
      selected_stn_count : Int;
      states : "Selectable Station States";
   END_VAR
   VAR CONSTANT
      initialize : String := 'initialize';
      all : String := 'all';
      non_hmi : String := 'non_hmi';
      hmi : String := 'hmi';
   END_VAR
BEGIN
   REGION "NOTES"
       (*
       The UDT containing all stations is too large to be instantiated in temp
       memory for this function. This is why you will see an initialization loop
       instead of a temp variable that gets returned later.
       *)
   END_REGION


   REGION "FOR ANY STATE"

       REGION "GET SELECTED STATION COUNT"
           #selected_stn_count := "Count Selected Stations"(#selected_stns.stns);
       END_REGION

       REGION "SELECTED STATION IS HMI"
           IF #selection_change.rising THEN
               #eval_station_is_hmi := "Is HMI Station"(#stns.stn[#selection_change.station_index]);
           END_IF;
           IF #selection_change.falling AND #selected_stn_count = 1 THEN
               #eval_station_is_hmi := "Is HMI Station"(#stns.stn["Get First Selected Station"(#selected_stns.stns)]);
           END_IF;
       END_REGION

   END_REGION


   REGION "SET STATE"

       REGION "ALL"
           // on first scan
           IF "FirstScan" THEN
               #states := "Set Selectable Station States"(#all);
           END_IF;
           // on selection change where last selected station is de-selected
           IF #selection_change.falling AND #selected_stn_count = 0 THEN
               #states := "Set Selectable Station States"(#all);
           END_IF;
       END_REGION

       REGION "NON HMI"
           // when no stations are selected and a non-hmi station is selected
           IF #selection_change.rising (*AND #selected_stn_count = 1*) THEN
               IF NOT #eval_station_is_hmi THEN
                   #states := "Set Selectable Station States"(#non_hmi);
               END_IF;
           END_IF;
       END_REGION

       REGION "HMI"
           // when no stations are selected and an hmi station is selected
           IF #selection_change.selection_change (*AND #selected_stn_count = 1*) THEN
               IF #eval_station_is_hmi THEN
                   #states := "Set Selectable Station States"(#hmi);
               END_IF;
           END_IF;
       END_REGION

   END_REGION


   REGION "ALL"
       IF #states.all THEN
           "Fill Int Array"(int_in := -1,
                        array_out => #selectable_stns);
           FOR #i := 0 TO "stnCount" DO
               #selectable_stns[#i] := #i;
           END_FOR;
           #selectable_stn_cnt := "stnCount";
       END_IF;
   END_REGION


   REGION "HMI & NON-HMI"
       IF #states.hmi OR #states.non_hmi THEN
           "Fill Int Array"(int_in := -1,
                        array_out => #selectable_stns);
           "Build HMI/Non-HMI List"(eval_stn_is_hmi := #eval_station_is_hmi,
                                    stns := #stns,
                                    selectable_stns := #selectable_stns,
                                    selectable_stn_count := #selectable_stn_cnt);
       END_IF;
   END_REGION


   REGION "HMI"
       IF #states.hmi THEN
           "Modify Selectable Station List: Matching WIP"(selection_change := #selection_change,
                                                          saved_wips := "HMI Stations: Saved Wips".stn,
                                                          selected_stations := #selected_stns,
                                                          selectable_stns := #selectable_stns,
                                                          selectable_stn_cnt := #selectable_stn_cnt,
                                                          visible_stations := #visible_stations);
       END_IF;
   END_REGION


   REGION "RETURN"
       (*
       Return values modified in "BUILD *" functions due to temp memory limit.
       *)
   END_REGION
END_FUNCTION

FUNCTION "Set Selectable Station States" : "Selectable Station States"   // FC107, SCL
{ S7_Optimized_Access := 'TRUE' }
VERSION : 0.1
   VAR_INPUT
      desired_state : String;
   END_VAR
   VAR_TEMP
      ret : "Selectable Station States";
   END_VAR
   VAR CONSTANT
      initialize : String := 'initialize';
      all : String := 'all';
      non_hmi : String := 'non_hmi';
      hmi : String := 'hmi';
   END_VAR
BEGIN
   REGION "SET ALL"
       IF #desired_state = #all THEN
           #ret.all := TRUE;
       END_IF;
   END_REGION


   REGION "SET NON_HMI"    
       IF #desired_state = #non_hmi THEN
           #ret.non_hmi := TRUE;
       END_IF;
   END_REGION


   REGION "SET HMI"
       IF #desired_state = #hmi THEN
           #ret.hmi := TRUE;
       END_IF;
   END_REGION


   REGION "RETURN"
       #"Set Selectable Station States" := #ret;
   END_REGION
END_FUNCTION

FUNCTION "Build HMI/Non-HMI List" : Void   // FC110, SCL
{ S7_Optimized_Access := 'TRUE' }
VERSION : 0.1
   VAR_INPUT
      eval_stn_is_hmi : Bool;
      stns : "Station: All Stations";
   END_VAR
   VAR_IN_OUT
      selectable_stns : Array[0.."stnCount"] of Int;
      selectable_stn_count : Int;
   END_VAR
   VAR_TEMP
      i : Int;
      t_selectable_stns : Array[0.."stnCount"] of Int;
      p_list : Int;
      this_stn_is_hmi : Bool;
   END_VAR
   VAR CONSTANT
      null_value : Int := -1;
   END_VAR
BEGIN
   REGION "NOTES"
       (*
       Checks to see if the evaluation station matches each station
       in the context of being or not being an HMI station.
       Returns the list of matching stations.
       *)
   END_REGION


   REGION "PREP LIST"
       "Fill Int Array"(int_in := #null_value,
                        array_out => #t_selectable_stns);
   END_REGION


   REGION "BUILD LIST"
       FOR #i := 0 TO "stnCount" DO
           #this_stn_is_hmi := "Is HMI Station"(#stns.stn[#i]);
           IF #eval_stn_is_hmi = #this_stn_is_hmi THEN
               #t_selectable_stns[#p_list] := #i;
               #p_list += 1;
           END_IF;
       END_FOR;
   END_REGION


   REGION "RETURN"
       #selectable_stns := #t_selectable_stns;
       #selectable_stn_count := #p_list;
   END_REGION
END_FUNCTION

